(* Logix 5000 project; controller Seperator 1756-L85E rev 34.11; software revision 34.00; part 2 of 7 *)
(* tags used below, declared in another part *)
   Inp : BOOL;   // Alarm Condition Input 1=Alarm
   Cfg_Exists : BOOL;   // 1=Alarm configured to exist, 0=Does not exist, don't scan
   Cfg_ResetReqd : BOOL;   // 1=Latched Alarm, a Reset is required to clear this Alarm
   Cfg_AckReqd : BOOL;   // 1=Acknowledge required for this Alarm
   Cfg_AllowShelve : BOOL;   // 1=Allow Operator to Shelve this Alarm
   Cfg_AllowDisable : BOOL;   // 1=Allow Maintenance to Disable this Alarm
   Cfg_Severity : SINT;   // Alarm Severity: 1=Low, 2=Medium, 3=High, 4=Highest
   Cfg_AlmMinOnT : DINT;   // Minimum time Alm output stays on (sec)
   Cfg_MaxShelfT : INT;   // Auto unshelve after shelved this long (1..32767 minutes)
   PCfg_AllowExist : BOOL;   // 1=Alarm can be configured to exist, 0=other configs make alarm meaningless
   PCmd_Ack : BOOL;   // Program Command to Acknowledge alarm
   PCmd_Suppress : BOOL;   // Program Command to Suppress by Design (inhibits new alarm)
   PCmd_Unsuppress : BOOL;   // Program Command to Unsuppress (allows new alarm)
   PCmd_Unshelve : BOOL;   // Program Command to Unshelve (e.g., on shift change)
   OCmd_Ack : BOOL;   // Operator Command to Acknowledge alarm
   OCmd_Shelve : BOOL;   // Operator Command to Shelve Alarm (inhibits new alarm)
   OCmd_Unshelve : BOOL;   // Operator Command to Unshelve alarm (allows new alarm)
   Alm : ALIAS FOR Com_AE.0;   // Alarm output 1=In Alarm
   Ack : ALIAS FOR Com_AE.1;   // Alarm acknowledged status: 1=Ack rcvd
   Shelved : ALIAS FOR Com_AE.3;   // 1=Alarm has been Shelved by Operator (inhibits new alarm)
   Suppressed : ALIAS FOR Com_AE.6;   // 1=Alarm has been Suppressed by Program (inhibits new alarm)
   Disabled : ALIAS FOR Com_AE.9;   // 1=Alarm has been Disabled by Maintanance (inhibits new alarm)
   P_Alarm : BOOL;   // Unique Parameter Name for auto - discovery
   Wrk_Suppressed : BOOL;   // Internal Alarm Suppressed Status
   Com_AE : INT;   // Communication with HMI / Alarm/Event Server (see bit descriptions)
   Starting : SFC_STEP;
   Stopped : SFC_STEP;
   Stopping : SFC_STEP;
(* P_Alarm, continued *)

ROUTINE Prescan   (* ladder *)
// Clear "lurking" Commands
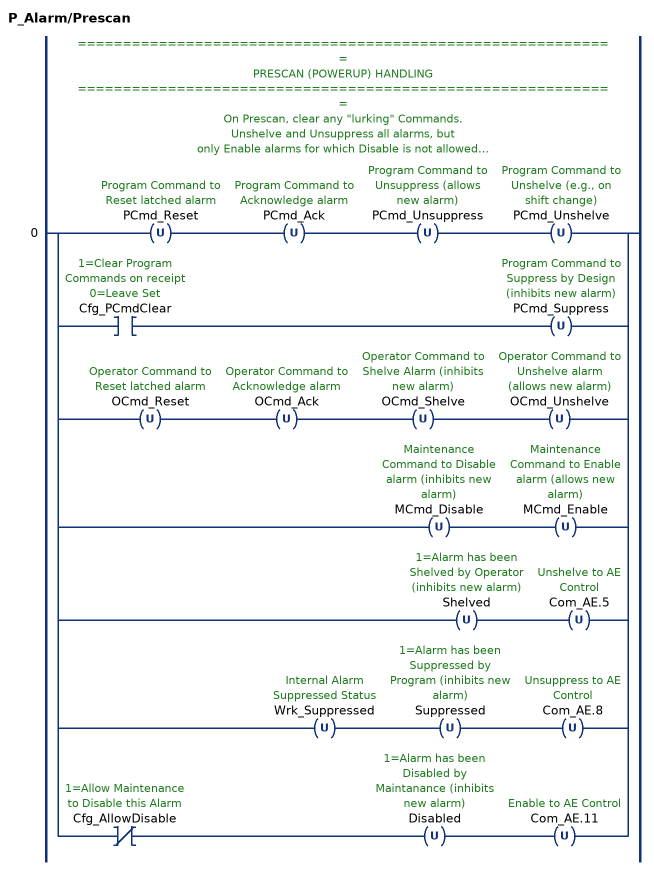
   // ============================================================
   // PRESCAN (POWERUP) HANDLING
   // ============================================================
   // On Prescan, clear any "lurking" Commands.
   // Unshelve and Unsuppress all alarms, but
   // only Enable alarms for which Disable is not allowed.
   // (Let Maintenance Disable persist through a power cycle...)
   // #####  V3.0-00  2013-06-30:  Added PCmd_Unshelve, AllowDisable, AllowShelve.  #####
   0: [OTU(PCmd_Reset) OTU(PCmd_Ack) OTU(PCmd_Unsuppress) OTU(PCmd_Unshelve) ,XIC(Cfg_PCmdClear) OTU(PCmd_Suppress) ,OTU(OCmd_Reset) OTU(OCmd_Ack) OTU(OCmd_Shelve) OTU(OCmd_Unshelve) ,OTU(MCmd_Disable) OTU(MCmd_Enable) ,OTU(Shelved) OTU(Com_AE.5) ,OTU(Wrk_Suppressed) OTU(Suppressed) OTU(Com_AE.8) ,XIO(Cfg_AllowDisable) OTU(Disabled) OTU(Com_AE.11) ];
END_ROUTINE
END_ADD_ON_INSTRUCTION

ADD_ON_INSTRUCTION P_Mode   (* revision 3.0 00 Release, vendor Rockwell Automation, ExecutePrescan, ExecuteEnableInFalse *)
// Mode
// Revision note:
// See Release Notes for Library version 3.0 for details on changes for this release. Containing objects MUST now expose OCmd_AcqLock and OCmd_Unlock. Made Operator Commands for going from Operator Locked to Program (unlocked) and Program (unlocked) to Operator Lock two-step processes.  Added Inf_Lib, Inf_Type.
// Help:
// Copyright © Rockwell Automation, Inc.  All Rights Reserved.
// This instruction provides selection of Mode (owner) for a Device level
// object  (from highest priority to lowest):
// *  No Mode (no owner, EnableIn is false)
// *  Hand (typically tracks hardwired control of device)
// *  Maint (Maintenance) (taken out of normal service for maintenance)
// *  Ovrd (Override) (typically used for process overrides)
// *  Prog  (Program) (automated control, and default if Cfg_ProgNorm = 1)
// *  Oper (Operator (manual control, and default if Cfg_ProgNorm = 0)
// (Program and Operator have the same priority.)
// The current mode is shown with Status bits and also as the primary
// Value for the instruction: an enumeration "Val" as follows:
//   0 = No Mode,
//   1 = Hand,
//   2 = Maintenance,
//   3 = Override,
//   4 = Program (Locked),
//   5 = Operator (Locked),
//   6 = Program (Unlocked, Oper default),
//   7 = Operator (Unlocked, Prog default),
//   8 = Program (Unlocked, = default),
//   9 = Operator (Unlocked, = default).
// When EnableIn is false, all ownership acquire/release and lock/unlock
// Commands are processed "behind the scenes", but the Mode is shown
// as "No Mode" (no owner).  When EnableIn becomes true, the Mode
// takes into account the Commands received -- in other words, the Mode
// becomes the one that would have been in effect had the EnableIn
// False / No Mode condition never occurred.
VAR_INPUT
   Inp_Hand : BOOL; {visible}   // 1=Acquire Hand (typ. hardwired local) Mode, 0=Release Hand Mode
   Inp_Ovrd : BOOL; {visible}   // 1=Acquire Override (higher priority program logic) Mode, 0=Release Override Mode
   Cfg_PCmdClear : BOOL := 1;   // 1=Clear Program Command on receipt; 0=Use Level-based (maintained) PCmds
   Cfg_OvrdOverLock : BOOL := 1;   // 1=Override supersedes Prog/Oper Lock, 0=don't override Lock
   Cfg_ProgDefault : BOOL;   // Default Mode: 1=Program Mode if no requests; 0=Operator Mode if no requests
   PCmd_Acq : BOOL;   // Program Command to Acquire Ownership (Oper to Prog)
   PCmd_Rel : BOOL;   // Program Command to Release Ownership (Prog to Oper)
   PCmd_Lock : BOOL;   // Program Command to Lock Mode in Prog
   PCmd_Unlock : BOOL;   // Program Command to Unlock Mode
   MCmd_Acq : BOOL;   // Maintenance Command to Acquire Ownership (Oper/Prog/Ovrd to Maint)
   MCmd_Rel : BOOL;   // Maintenance Command to Release Ownership (Maint to Oper/Prog/Ovrd)
   OCmd_AcqLock : BOOL;   // Operator Command to Acquire (Prog to Oper) / Lock Ownership
   OCmd_UnlockRel : BOOL;   // Operator Command to Unlock / Release (Oper to Prog) Ownership
END_VAR
VAR_OUTPUT
   Val : DINT; {access Read Only}   // Mode enum: 0=No, 1=H, 2=M, 3=!, 4=P Lock, 5=O Lock, 6=P (O Def), 7=O (P Def), 8=P (= Def), 9=O (= Def)
   Sts_Hand : BOOL; {access Read Only, visible}   // 1=Mode is Hand (supersedes Maint, Ovrd, Prog, Oper)
   Sts_Maint : BOOL; {access Read Only, visible}   // 1=Mode is Maintenance (supersedes Ovrd, Prog, Oper)
   Sts_Ovrd : BOOL; {access Read Only, visible}   // 1=Mode is Override (supersedes Prog, Oper)
   Sts_Prog : BOOL; {access Read Only, visible}   // 1=Mode is Program
   Sts_Oper : BOOL := 1; {access Read Only, visible}   // 1=Mode is Operator
   Sts_ProgOperLock : BOOL; {access Read Only, visible}   // 1=Program or Operator has requested Mode Lock
   Sts_ProgOperSel : BOOL; {access Read Only}   // Prog/Oper selection 1=Program, 0=Operator
   Sts_NoMode : BOOL; {access Read Only}   // 1=Mode is No Mode (no owner, disabled or not scanned)
   Rdy_MAcq : BOOL; {access Read Only}   // 1=Ready for MCmd_Acq, enable button
   Rdy_MRel : BOOL; {access Read Only}   // 1=Ready for MCmd_Rel, enable button
   Rdy_OAcq : BOOL; {access Read Only}   // 1=Ready for OCmd_AcqLock, enable Acquire (to Oper) button
   Rdy_OLock : BOOL; {access Read Only}   // 1=Ready for OCmd_AcqLock, enable Oper Lock button
   Rdy_OUnlock : BOOL; {access Read Only}   // 1=Ready for OCmd_UnlockRel, enable Oper Unlock button
   Rdy_ORel : BOOL; {access Read Only}   // 1=Ready for OCmd_UnlockRel, enable Release (to Prog) button
   P_Mode : BOOL;   // Unique Parameter Name for auto - discovery
END_VAR
VAR
   Wrk_Locked : BOOL; {access None}   // 1=Program/Operator Mode selection is Locked
   Wrk_Prog : BOOL; {access None}   // Internal Program (1) / Operator (0) Mode selection
   Wrk_Maint : BOOL; {access None}   // Internal Maintenance Mode
   Inf_Lib : STRING_12 := 'RA-BAS'; {access Read Only}   // Display Library for Faceplate call-up
   Inf_Type : STRING_16_UDT := 'P_Mode'; {access Read Only}   // Must contain AOI name, used for HMI and Information S/W
END_VAR

ROUTINE EnableInFalse   (* ladder *)
// Processes received Commands, but shows "NO mode" (no owner)
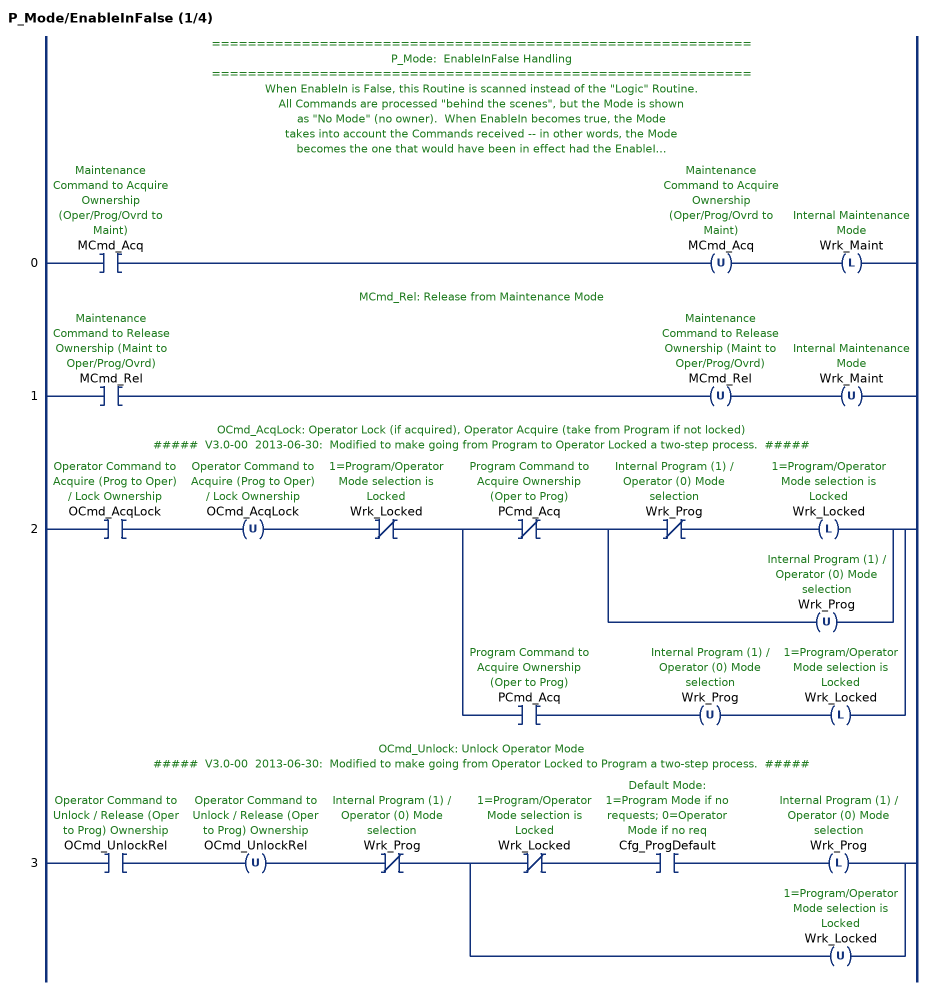
   // ============================================================
   // P_Mode:  EnableInFalse Handling
   // ============================================================
   // When EnableIn is False, this Routine is scanned instead of the "Logic" Routine.
   // All Commands are processed "behind the scenes", but the Mode is shown
   // as "No Mode" (no owner).  When EnableIn becomes true, the Mode
   // takes into account the Commands received -- in other words, the Mode
   // becomes the one that would have been in effect had the EnableIn
   // False / No Mode condition never occurred.
   // ============================================================
   // COMMAND HANDLING
   // ============================================================
   // NOTE:  These rungs MUST be in the order given to meet the following
   // multiple-actions-at-the-same-time scenarios:
   // * Maintenance Release beats Maintenance Acquire
   // * Program Release beats Program Acquire
   // * Program Unlock beats Program Lock
   // * Operator Unlock beats Operator Acquire and Lock (results in Oper Unlocked)
   // * Operator Acquire/Lock must come after Program Unlock
   // * Program Acquire must come after Operator Unlock
   // ============================================================
   // MCmd_Acq: Acquire for Maintenance Mode
   0: XIC(MCmd_Acq)OTU(MCmd_Acq)OTL(Wrk_Maint);
   // MCmd_Rel: Release from Maintenance Mode
   1: XIC(MCmd_Rel)OTU(MCmd_Rel)OTU(Wrk_Maint);
   // OCmd_AcqLock: Operator Lock (if acquired), Operator Acquire (take from Program if not locked)
   // #####  V3.0-00  2013-06-30:  Modified to make going from Program to Operator Locked a two-step process.  #####
   2: XIC(OCmd_AcqLock)OTU(OCmd_AcqLock)XIO(Wrk_Locked)[XIO(PCmd_Acq) [XIO(Wrk_Prog) OTL(Wrk_Locked) ,OTU(Wrk_Prog) ] ,XIC(PCmd_Acq) OTU(Wrk_Prog) OTL(Wrk_Locked) ];
   // OCmd_Unlock: Unlock Operator Mode
   // #####  V3.0-00  2013-06-30:  Modified to make going from Operator Locked to Program a two-step process.  #####
   3: XIC(OCmd_UnlockRel)OTU(OCmd_UnlockRel)XIO(Wrk_Prog)[XIO(Wrk_Locked) XIC(Cfg_ProgDefault) OTL(Wrk_Prog) ,OTU(Wrk_Locked) ];
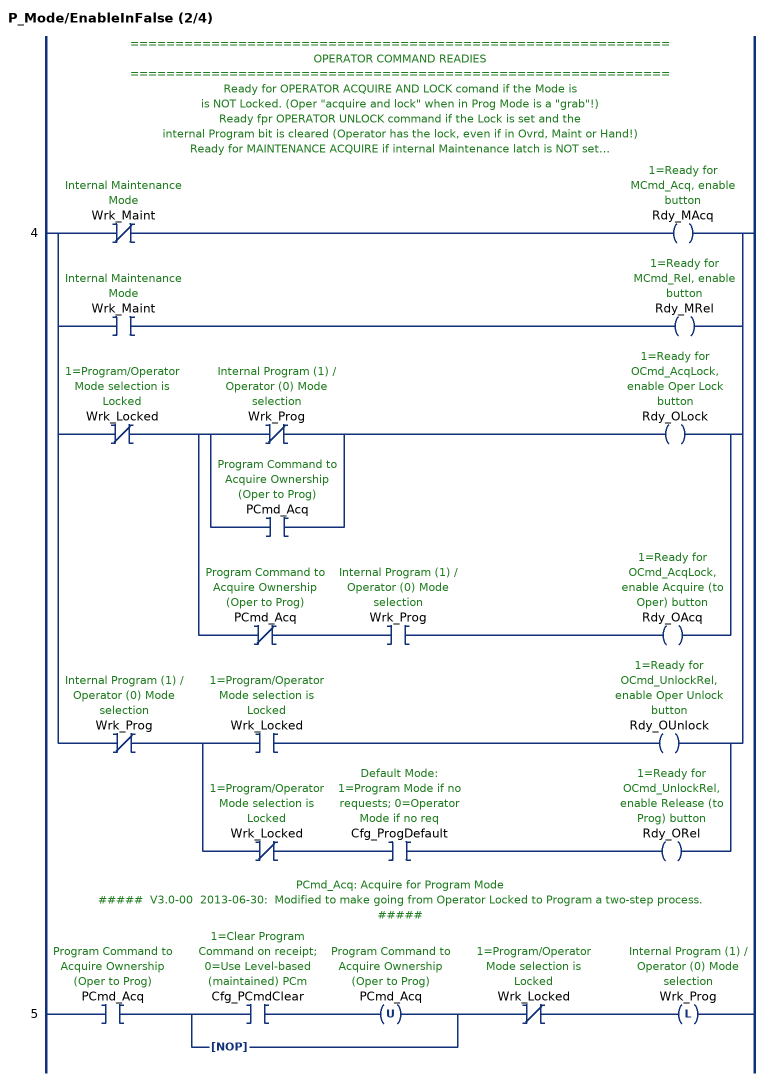
   // ============================================================
   // OPERATOR COMMAND READIES
   // ============================================================
   // Ready for OPERATOR ACQUIRE AND LOCK comand if the Mode is
   //  is NOT Locked. (Oper "acquire and lock" when in Prog Mode is a "grab"!)
   // Ready fpr OPERATOR UNLOCK command if the Lock is set and the
   // internal Program bit is cleared (Operator has the lock, even if in Ovrd, Maint or Hand!)
   // Ready for MAINTENANCE ACQUIRE if internal Maintenance latch is NOT set.
   // Ready for MAINTENANCE RELEASE if internal Maintenance latch IS set.
   // #####  V3.0-00  2013-06-30:  Modified Rdy_Unlock for two-step Operator Locked to Program process.  #####
   4: [XIO(Wrk_Maint) OTE(Rdy_MAcq) ,XIC(Wrk_Maint) OTE(Rdy_MRel) ,XIO(Wrk_Locked) [[XIO(Wrk_Prog) ,XIC(PCmd_Acq) ] OTE(Rdy_OLock) ,XIO(PCmd_Acq) XIC(Wrk_Prog) OTE(Rdy_OAcq) ] ,XIO(Wrk_Prog) [XIC(Wrk_Locked) OTE(Rdy_OUnlock) ,XIO(Wrk_Locked) XIC(Cfg_ProgDefault) OTE(Rdy_ORel) ] ];
   // PCmd_Acq: Acquire for Program Mode
   // #####  V3.0-00  2013-06-30:  Modified to make going from Operator Locked to Program a two-step process.  #####
   5: XIC(PCmd_Acq)[XIC(Cfg_PCmdClear) OTU(PCmd_Acq) ,NOP() ]XIO(Wrk_Locked)OTL(Wrk_Prog);
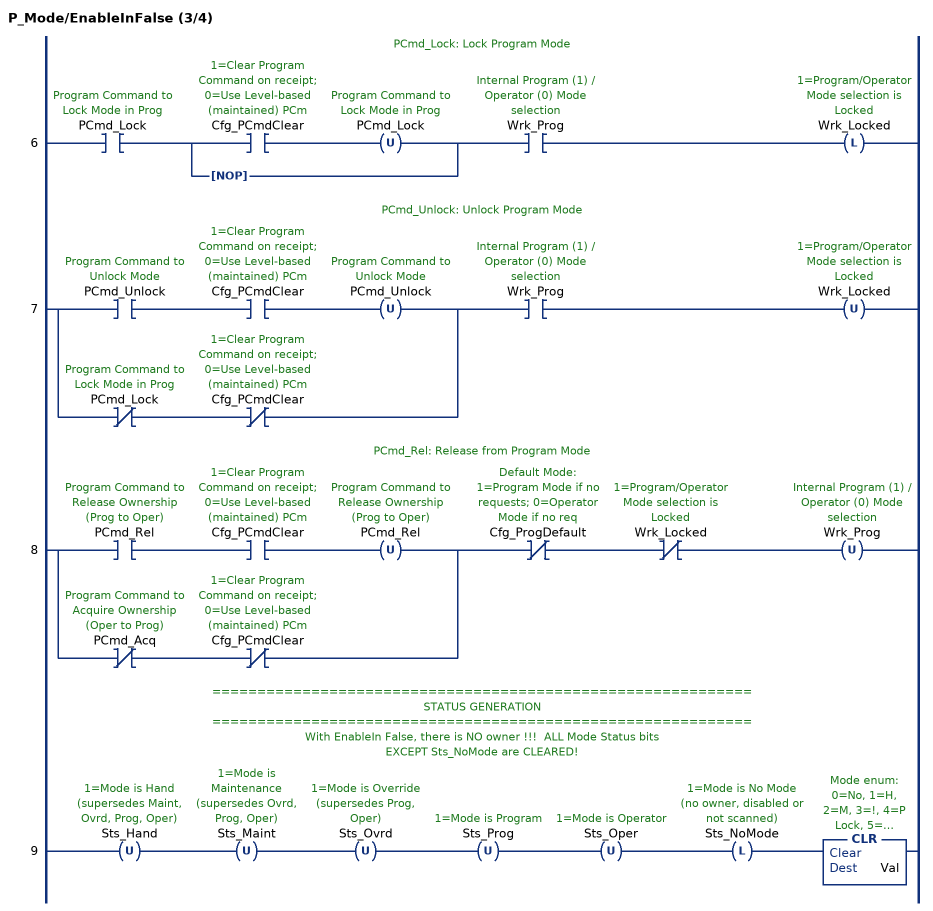
   // PCmd_Lock: Lock Program Mode
   6: XIC(PCmd_Lock)[XIC(Cfg_PCmdClear) OTU(PCmd_Lock) ,NOP() ]XIC(Wrk_Prog)OTL(Wrk_Locked);
   // PCmd_Unlock: Unlock Program Mode
   7: [XIC(PCmd_Unlock) XIC(Cfg_PCmdClear) OTU(PCmd_Unlock) ,XIO(PCmd_Lock) XIO(Cfg_PCmdClear) ]XIC(Wrk_Prog)OTU(Wrk_Locked);
   // PCmd_Rel: Release from Program Mode
   8: [XIC(PCmd_Rel) XIC(Cfg_PCmdClear) OTU(PCmd_Rel) ,XIO(PCmd_Acq) XIO(Cfg_PCmdClear) ]XIO(Cfg_ProgDefault)XIO(Wrk_Locked)OTU(Wrk_Prog);
   // ============================================================
   // STATUS GENERATION
   // ============================================================
   // With EnableIn False, there is NO owner !!!  ALL Mode Status bits
   // EXCEPT Sts_NoMode are CLEARED!
   9: OTU(Sts_Hand)OTU(Sts_Maint)OTU(Sts_Ovrd)OTU(Sts_Prog)OTU(Sts_Oper)OTL(Sts_NoMode)CLR(Val);
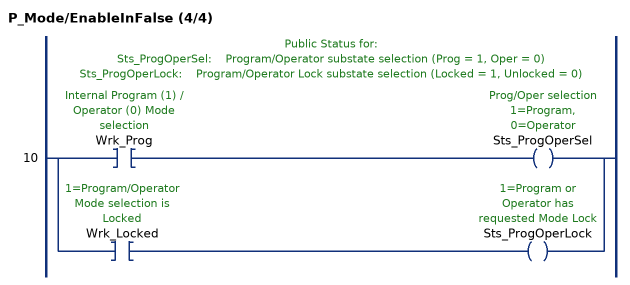
   // Public Status for:
   // Sts_ProgOperSel:    Program/Operator substate selection (Prog = 1, Oper = 0)
   // Sts_ProgOperLock:    Program/Operator Lock substate selection (Locked = 1, Unlocked = 0)
   10: [XIC(Wrk_Prog) OTE(Sts_ProgOperSel) ,XIC(Wrk_Locked) OTE(Sts_ProgOperLock) ];
END_ROUTINE

ROUTINE Logic   (* ladder *)
// Selects Modes (Hand, Maint, Ovrd, Oper, Prog) based on Inputs and Commands
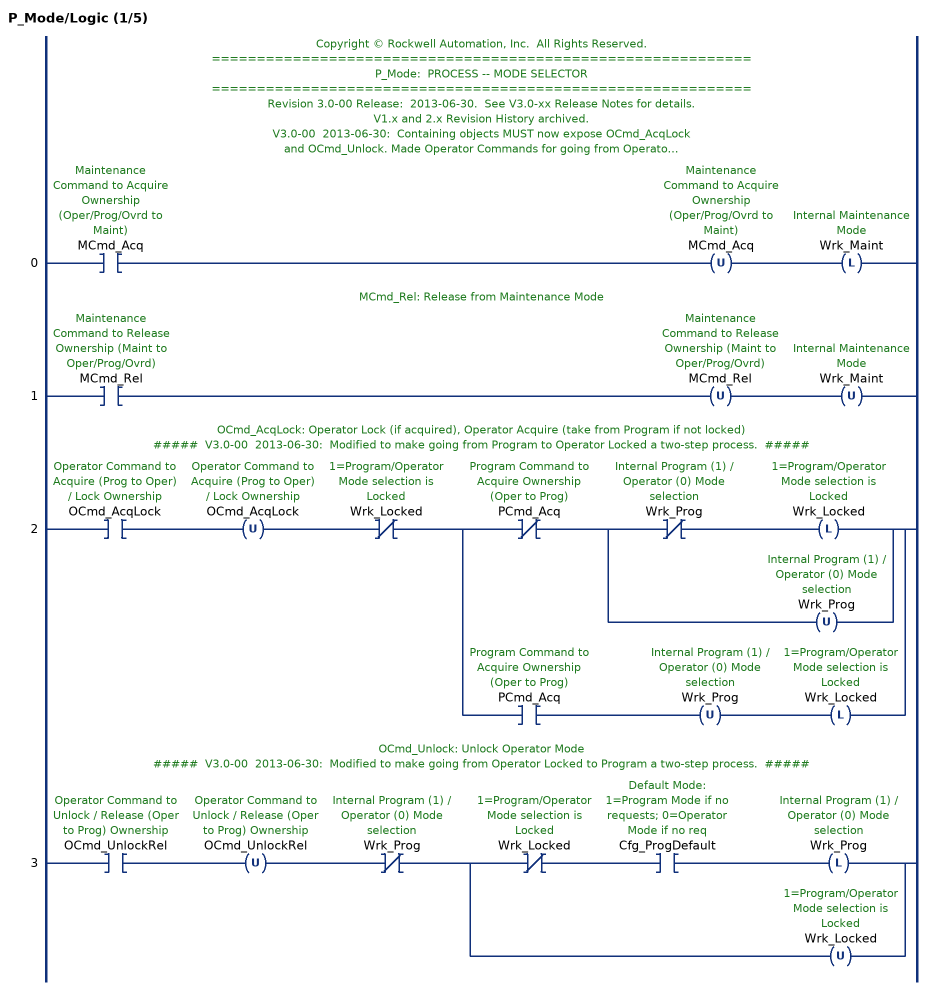
   // Copyright © Rockwell Automation, Inc.  All Rights Reserved.
   // ============================================================
   // P_Mode:  PROCESS -- MODE SELECTOR
   // ============================================================
   // Revision 3.0-00 Release:  2013-06-30.  See V3.0-xx Release Notes for details.
   // V1.x and 2.x Revision History archived.
   // V3.0-00  2013-06-30:  Containing objects MUST now expose OCmd_AcqLock
   // and OCmd_Unlock. Made Operator Commands for going from Operator
   // Locked to Program (unlocked) and Program (unlocked) to Operator
   // Lock two-step processes.  Added Inf_Lib, Inf_Type.
   // ============================================================
   // This instruction provides selection of Mode (owner) for a Device level
   // object  (from highest priority to lowest):
   // * NO Mode (EnableIn is false)
   // *  Hand (typically tracks hardwired control of device)
   // *  Maint (Maintenance) (taken out of normal service for maintenance)
   // *  Ovrd (Override) (typically used for process overrides)
   // *  Prog  (Program) (automated control, and default if Cfg_ProgNorm = 1)
   // *  Oper (Operator (manual control, and default if Cfg_ProgNorm = 0)
   // The current mode is shown with Status bits and also as the
   // primary Value for the instruction: an enumeration as follows:
   // 0 = No Mode, 1 = Hand, 2 = Maintenance, 3 = Override,
   // 4 = Program (Locked), 5 = Operator (Locked),
   // 6 = Program (Unlocked, Oper default), 7 = Operator (Unlocked, Prog default),
   // 8 = Program (Unlocked, Prog default), 9 = Operator (Unlocked, Oper default).
   // ============================================================
   // COMMAND HANDLING
   // ============================================================
   // NOTE:  These rungs MUST be in the order given to meet the following
   // multiple-actions-at-the-same-time scenarios:
   // * Maintenance Release beats Maintenance Acquire
   // * Program Release beats Program Acquire
   // * Program Unlock beats Program Lock
   // * Operator Unlock beats Operator Acquire / Lock (results in Oper Unlocked)
   // * Program Acquire must come after Operator Unlock
   // If Cfg_ProgDefault = 1, the Mode defaults to Program
   // (instead of Operator) if all other Modes release their requests.
   // ============================================================
   // MCmd_Acq: Acquire for Maintenance Mode
   0: XIC(MCmd_Acq)OTU(MCmd_Acq)OTL(Wrk_Maint);
   // MCmd_Rel: Release from Maintenance Mode
   1: XIC(MCmd_Rel)OTU(MCmd_Rel)OTU(Wrk_Maint);
   // OCmd_AcqLock: Operator Lock (if acquired), Operator Acquire (take from Program if not locked)
   // #####  V3.0-00  2013-06-30:  Modified to make going from Program to Operator Locked a two-step process.  #####
   2: XIC(OCmd_AcqLock)OTU(OCmd_AcqLock)XIO(Wrk_Locked)[XIO(PCmd_Acq) [XIO(Wrk_Prog) OTL(Wrk_Locked) ,OTU(Wrk_Prog) ] ,XIC(PCmd_Acq) OTU(Wrk_Prog) OTL(Wrk_Locked) ];
   // OCmd_Unlock: Unlock Operator Mode
   // #####  V3.0-00  2013-06-30:  Modified to make going from Operator Locked to Program a two-step process.  #####
   3: XIC(OCmd_UnlockRel)OTU(OCmd_UnlockRel)XIO(Wrk_Prog)[XIO(Wrk_Locked) XIC(Cfg_ProgDefault) OTL(Wrk_Prog) ,OTU(Wrk_Locked) ];
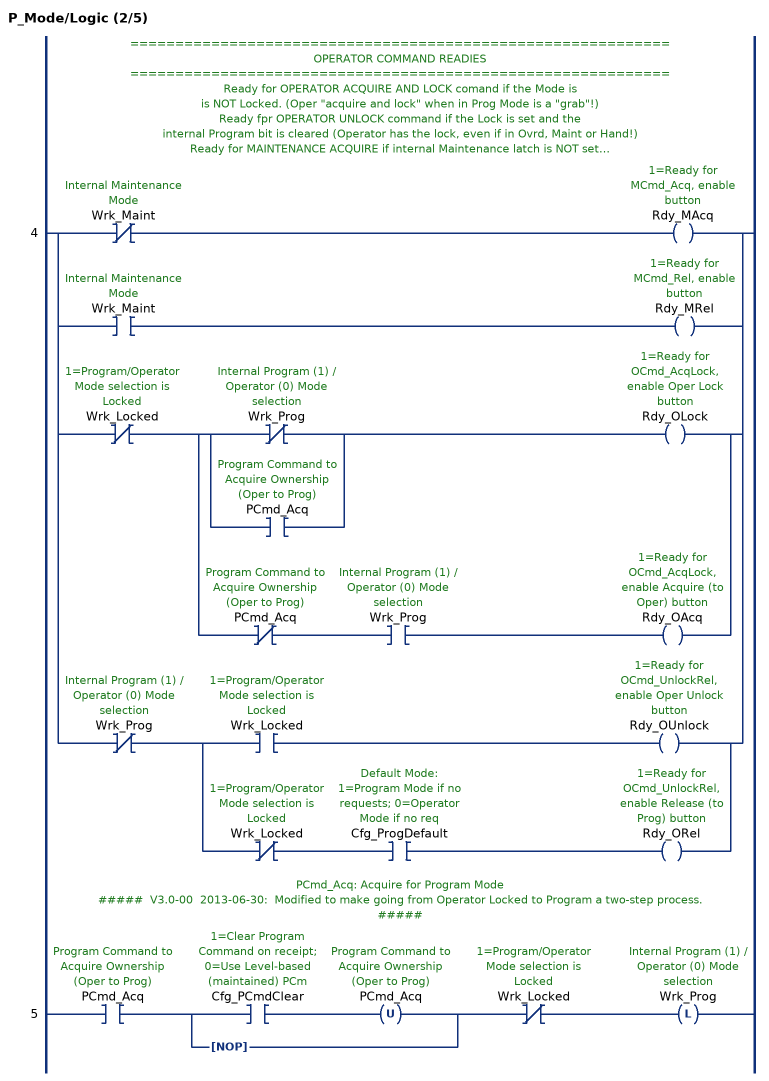
   // ============================================================
   // OPERATOR COMMAND READIES
   // ============================================================
   // Ready for OPERATOR ACQUIRE AND LOCK comand if the Mode is
   //  is NOT Locked. (Oper "acquire and lock" when in Prog Mode is a "grab"!)
   // Ready fpr OPERATOR UNLOCK command if the Lock is set and the
   // internal Program bit is cleared (Operator has the lock, even if in Ovrd, Maint or Hand!)
   // Ready for MAINTENANCE ACQUIRE if internal Maintenance latch is NOT set.
   // Ready for MAINTENANCE RELEASE if internal Maintenance latch IS set.
   // #####  V3.0-00  2013-06-30:  Modified Rdy_Unlock for two-step Operator Locked to Program process.  #####
   4: [XIO(Wrk_Maint) OTE(Rdy_MAcq) ,XIC(Wrk_Maint) OTE(Rdy_MRel) ,XIO(Wrk_Locked) [[XIO(Wrk_Prog) ,XIC(PCmd_Acq) ] OTE(Rdy_OLock) ,XIO(PCmd_Acq) XIC(Wrk_Prog) OTE(Rdy_OAcq) ] ,XIO(Wrk_Prog) [XIC(Wrk_Locked) OTE(Rdy_OUnlock) ,XIO(Wrk_Locked) XIC(Cfg_ProgDefault) OTE(Rdy_ORel) ] ];
   // PCmd_Acq: Acquire for Program Mode
   // #####  V3.0-00  2013-06-30:  Modified to make going from Operator Locked to Program a two-step process.  #####
   5: XIC(PCmd_Acq)[XIC(Cfg_PCmdClear) OTU(PCmd_Acq) ,NOP() ]XIO(Wrk_Locked)OTL(Wrk_Prog);
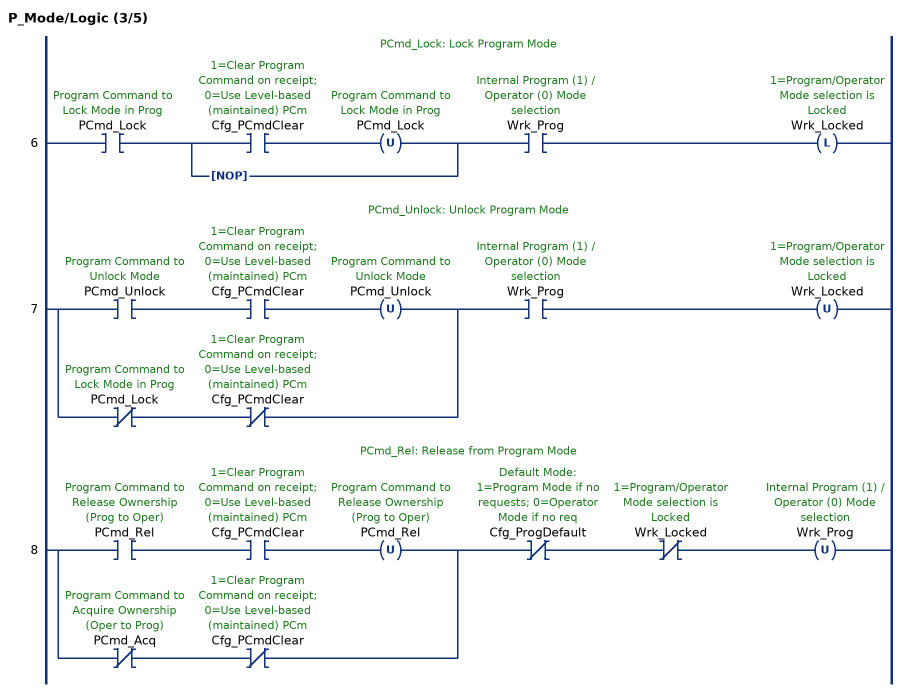
   // PCmd_Lock: Lock Program Mode
   6: XIC(PCmd_Lock)[XIC(Cfg_PCmdClear) OTU(PCmd_Lock) ,NOP() ]XIC(Wrk_Prog)OTL(Wrk_Locked);
   // PCmd_Unlock: Unlock Program Mode
   7: [XIC(PCmd_Unlock) XIC(Cfg_PCmdClear) OTU(PCmd_Unlock) ,XIO(PCmd_Lock) XIO(Cfg_PCmdClear) ]XIC(Wrk_Prog)OTU(Wrk_Locked);
   // PCmd_Rel: Release from Program Mode
   8: [XIC(PCmd_Rel) XIC(Cfg_PCmdClear) OTU(PCmd_Rel) ,XIO(PCmd_Acq) XIO(Cfg_PCmdClear) ]XIO(Cfg_ProgDefault)XIO(Wrk_Locked)OTU(Wrk_Prog);
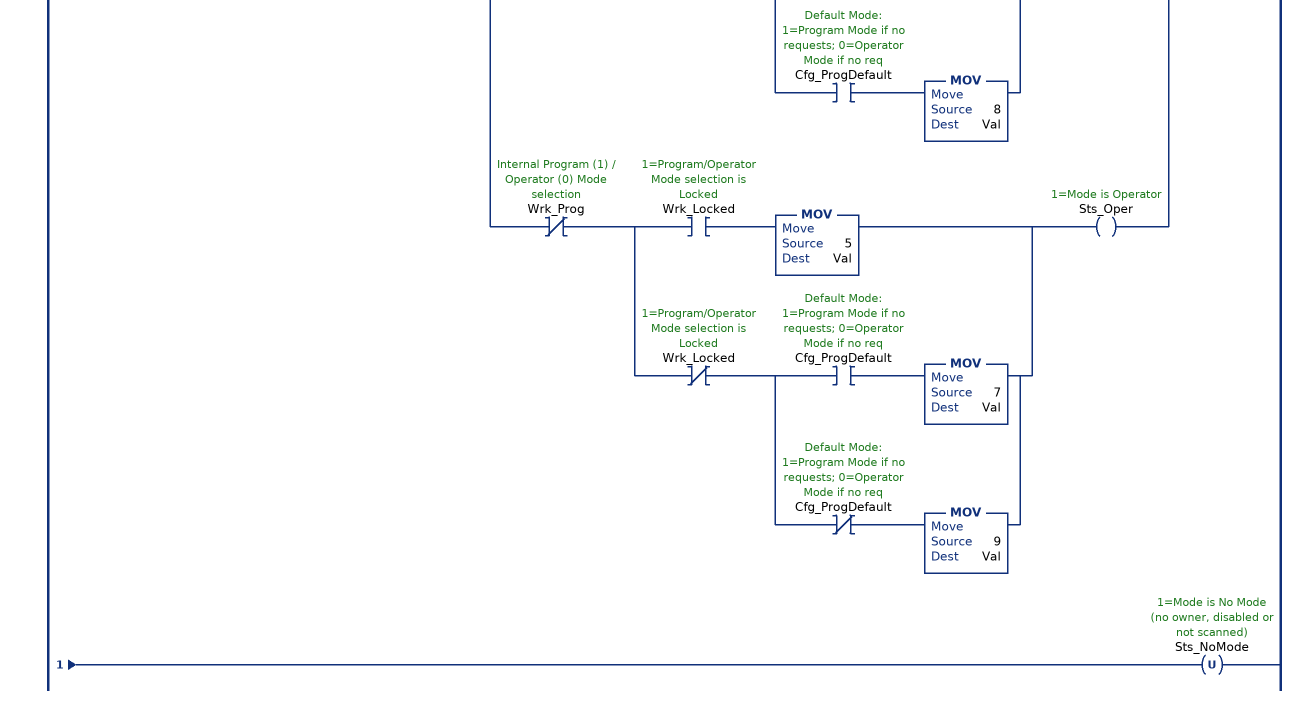
   // ============================================================
   // STATUS GENERATION
   // ============================================================
   // This rung determines the Mode based on the states of the inputs and internal working bits.
   // The logic here does the vast mahority of the implementation of the Mode selection rules.
   // Between the internal working bits used above and the rules implemented here,
   // outside objects cannot manipulate the state of this object by setting/clearing its Status bits.
   // Public Status is generated for:
   // *  Hand Mode
   // *  Maintenance Mode
   // *  Override Mode
   // *  Program Mode
   // *  Operator Mode
   // *  No Mode (none of the above)
   9: [XIC(Inp_Hand) OTE(Sts_Hand) MOV(1,Val) ,XIO(Inp_Hand) [XIC(Wrk_Maint) OTE(Sts_Maint) MOV(2,Val) ,XIO(Wrk_Maint) [XIC(Inp_Ovrd) [XIO(Wrk_Locked) ,XIC(Cfg_OvrdOverLock) ,XIC(Sts_Ovrd) ] OTE(Sts_Ovrd) MOV(3,Val) ,XIO(Sts_Ovrd) [XIC(Wrk_Prog) [XIC(Wrk_Locked) MOV(4,Val) ,XIO(Wrk_Locked) [XIO(Cfg_ProgDefault) MOV(6,Val) ,XIC(Cfg_ProgDefault) MOV(8,Val) ] ] OTE(Sts_Prog) ,XIO(Wrk_Prog) [XIC(Wrk_Locked) MOV(5,Val) ,XIO(Wrk_Locked) [XIC(Cfg_ProgDefault) MOV(7,Val) ,XIO(Cfg_ProgDefault) MOV(9,Val) ] ] OTE(Sts_Oper) ] ] ] ]OTU(Sts_NoMode);
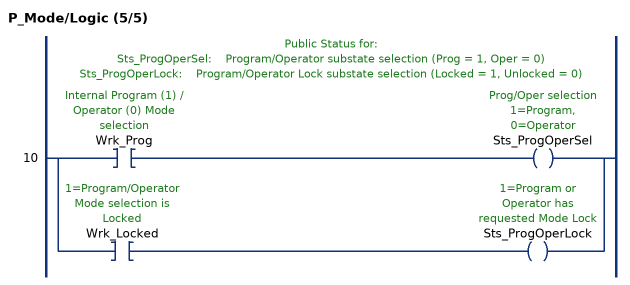
   // Public Status for:
   // Sts_ProgOperSel:    Program/Operator substate selection (Prog = 1, Oper = 0)
   // Sts_ProgOperLock:    Program/Operator Lock substate selection (Locked = 1, Unlocked = 0)
   10: [XIC(Wrk_Prog) OTE(Sts_ProgOperSel) ,XIC(Wrk_Locked) OTE(Sts_ProgOperLock) ];
END_ROUTINE

ROUTINE Prescan   (* ladder *)
// Clear "lurking" Commands
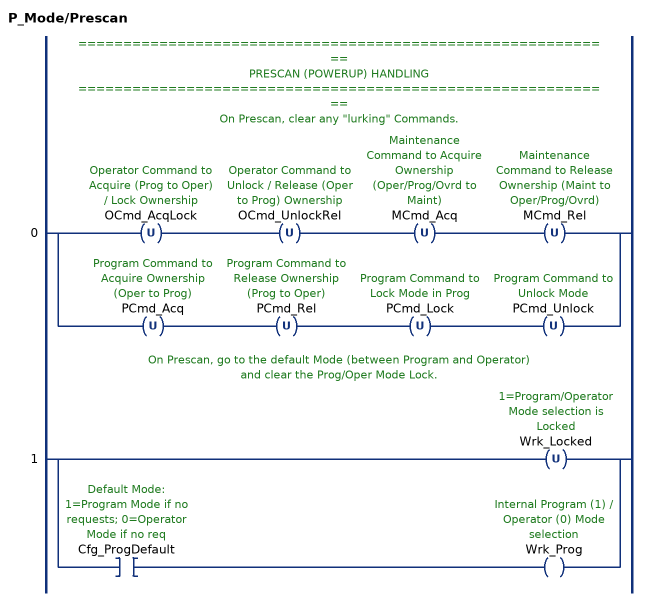
   // ============================================================
   // PRESCAN (POWERUP) HANDLING
   // ============================================================
   // On Prescan, clear any "lurking" Commands.
   0: [OTU(OCmd_AcqLock) OTU(OCmd_UnlockRel) OTU(MCmd_Acq) OTU(MCmd_Rel) ,OTU(PCmd_Acq) OTU(PCmd_Rel) OTU(PCmd_Lock) OTU(PCmd_Unlock) ];
   // On Prescan, go to the default Mode (between Program and Operator)
   // and clear the Prog/Oper Mode Lock.
   1: [OTU(Wrk_Locked) ,XIC(Cfg_ProgDefault) OTE(Wrk_Prog) ];
END_ROUTINE
END_ADD_ON_INSTRUCTION

ADD_ON_INSTRUCTION P_Motor   (* revision 3.0 04 Release, vendor Rockwell Automation, ExecutePrescan, ExecuteEnableInFalse *)
// Single Speed Motor
// Revision note:
// See Release Notes for Library version 3.0 for details on changes for this release. Corrected Parameter descriptions and default configuration values for alarms only.
// Help:
// Copyright © Rockwell Automation, Inc.  All Rights Reserved.
// This Instruction controls and monitors a single-speed motor
// (FVNR, soft-start, etc.) and provides:
// *  Monitoring of run feedback, display of actual motor status
// *  Detection of Failure to Start, Failure to Stop
// *  Monitoring of a Permissive condition to allow starting
// *  Monitoring of an Interlock condition to stop / prevent starting
// *  Simulation, providing feedback of a working motor while disabling outputs
// *  Monitoring of I/O communication faults
// *  Alarms for Fail to Start, Fail to Stop, Interlock Trip, I/O Fault
// *  Options to shed (stop motor) on Fail to Start or I/O Fault
// *  Operation in Hand, Maintenance, Override, Program and Operator Modes
// *  Option to automatically reset faults and alarms when operator commands
//      motor to start or stop
// *  Supports HMI "breadcrumbs" for Alarm Inhibited, Bad Configuration,
//      Not Ready, Maintenance Bypass Active
// *  "Available" status for use by automation logic to know whether motor
//      can be controlled by other objects.
// Modes are provided by a P_Mode AOI instance.
// Alarms are provided by P_Alarm AOI instances.
// Modes of operation: Operator, Program, Override, Maintenance, Hand
VAR_INPUT
   Inp_RunFdbk : BOOL; {visible}   // Input Signal: RUN feedback from motor
   Inp_PermOK : BOOL := 1; {visible}   // 1=Permissives OK, motor can start
   Inp_NBPermOK : BOOL := 1; {visible}   // 1=Non-Bypassable Permissives OK, motor can start
   Inp_IntlkOK : BOOL := 1; {visible}   // 1=Interlocks OK, motor can start/run
   Inp_NBIntlkOK : BOOL := 1; {visible}   // 1=Non-Bypassable Interlocks OK, motor can start/run
   Inp_IOFault : BOOL;   // Input Communication Status 0=OK, 1=fail
   Inp_Sim : BOOL;   // 1=Simulate working motor; 0=Start/Stop/ Monitor actual motor
   Inp_Hand : ALIAS FOR Mode.Inp_Hand;
   Inp_Ovrd : ALIAS FOR Mode.Inp_Ovrd;
   Inp_OvrdCmd : DINT;   // Override Mode Command: 0=None, 1=Stop, 2=Start
   Inp_Reset : BOOL;   // 1=Reset all fault conditions and latched Alarms
   Cfg_HasRunFdbk : BOOL;   // 1=Motor provides run feedback
   Cfg_UseRunFdbk : BOOL;   // 1=Motor run feedback should be used for failure checking
   Cfg_AllowLocal : BOOL;   // 1=Allow Local Start/Stop without alarm, 0=Start/Stop from HMI/prog only
   Cfg_HasPermObj : BOOL;   // 1=Enable navigation to permissive object
   Cfg_HasIntlkObj : BOOL;   // 1=Enable navigation to interlock object
   Cfg_HasResInhObj : BOOL;   // 1=Enable navigation to restart inhibit object
   Cfg_HasRunTimeObj : BOOL;   // 1=Enable navigation to run time object
   Cfg_HasOvldObj : BOOL;   // 1=Enable navigation to overload object
   Cfg_PCmdClear : ALIAS FOR Mode.Cfg_PCmdClear;
   Cfg_ProgDefault : ALIAS FOR Mode.Cfg_ProgDefault;
   Cfg_OperStopPrio : BOOL;   // 1=OCmd_Stop available in any mode, 0=OCmd_Stop only in Oper, Maint modes.
   Cfg_OCmdResets : BOOL;   // 1=New Oper motor cmd. resets fault, 0=reset req'd to clear fault
   Cfg_OvrdPermIntlk : BOOL;   // 1=Override ignores Bypassable Perm/ Intlk; 0=always use Perm/Intlk
   Cfg_ShedOnFailToStart : BOOL := 1;   // 1=Stop Motor and Alarm on Fail to Start; 0=Alarm only on Fail to Start
   Cfg_ShedOnIOFault : BOOL := 1;   // 1=Stop Motor and Alarm on I/O Fault; 0=Alarm only on I/O Fault
   Cfg_HasFailToStartAlm : ALIAS FOR FailToStart.Cfg_Exists;   // 1=Fail to Start Alarm exists and will be checked
   Cfg_HasFailToStopAlm : ALIAS FOR FailToStop.Cfg_Exists;   // 1=Fail to Stop Alarm exists and will be checked
   Cfg_HasIntlkTripAlm : ALIAS FOR IntlkTrip.Cfg_Exists;   // 1=Interlock Trip Alarm exists and will be checked
   Cfg_HasIOFaultAlm : ALIAS FOR IOFault.Cfg_Exists;   // 1=I/O Fault Alarm exists and will be checked
   Cfg_FailToStartResetReqd : ALIAS FOR FailToStart.Cfg_ResetReqd;   // 1=Reset required to clear Fail to Start Alarm
   Cfg_FailToStopResetReqd : ALIAS FOR FailToStop.Cfg_ResetReqd;   // 1=Reset required to clear Fail to Stop Alarm
   Cfg_IntlkTripResetReqd : ALIAS FOR IntlkTrip.Cfg_ResetReqd;   // 1=Reset required to clear Interlock Trip Alarm
   Cfg_IOFaultResetReqd : ALIAS FOR IOFault.Cfg_ResetReqd;   // 1=Reset required to clear I/O Fault Alarm
   Cfg_FailToStartAckReqd : ALIAS FOR FailToStart.Cfg_AckReqd;   // 1=Acknowledge required for Fail to Start Alarm
   Cfg_FailToStopAckReqd : ALIAS FOR FailToStop.Cfg_AckReqd;   // 1=Acknowledge required for Fail to Stop Alarm
   Cfg_IntlkTripAckReqd : ALIAS FOR IntlkTrip.Cfg_AckReqd;   // 1=Acknowledge required for Interlock Trip Alarm
   Cfg_IOFaultAckReqd : ALIAS FOR IOFault.Cfg_AckReqd;   // 1=Acknowledge required for I/O Fault Alarm
   Cfg_FailToStartSeverity : ALIAS FOR FailToStart.Cfg_Severity;   // Fail To Start Alarm Severity: 1=low, 2=medium, 3=high, 4=highest
   Cfg_FailToStopSeverity : ALIAS FOR FailToStop.Cfg_Severity;   // Fail To Stop Alarm Severity: 1=low, 2=medium, 3=high, 4=highest
   Cfg_IntlkTripSeverity : ALIAS FOR IntlkTrip.Cfg_Severity;   // Interlock Trip Alarm Severity: 1=low, 2=medium, 3=high, 4=highest
   Cfg_IOFaultSeverity : ALIAS FOR IOFault.Cfg_Severity;   // I/O Fault Alarm Severity: 1=low, 2=medium, 3=high, 4=highest
   Cfg_SimFdbkT : DINT := 2;   // Feedback delay in Simulation (sec)
   Cfg_FailToStartT : DINT := 10;   // Time after Start for running feedback before Fault (sec)
   Cfg_FailToStopT : DINT := 10;   // Time after Stop for stopped feedback (=0) before Fault (sec)
   PSet_Owner : DINT;   // Program Owner Request ID (non-zero) or Release (zero)
   PCmd_Start : BOOL;   // Program Command to Start Motor
   PCmd_Stop : BOOL;   // Program Command to Stop Motor
   PCmd_Acq : ALIAS FOR Mode.PCmd_Acq;
   PCmd_Rel : ALIAS FOR Mode.PCmd_Rel;
   PCmd_Lock : ALIAS FOR Mode.PCmd_Lock;
   PCmd_Unlock : ALIAS FOR Mode.PCmd_Unlock;
   PCmd_Reset : BOOL;   // Program Command to Reset all Alarms requiring Reset
   PCmd_FailToStartAck : ALIAS FOR FailToStart.PCmd_Ack;   // Program Command to Acknowledge Fail to Start Alarm
   PCmd_FailToStartSuppress : ALIAS FOR FailToStart.PCmd_Suppress;   // Program Command to Suppress Fail to Start Alarm
   PCmd_FailToStartUnsuppress : ALIAS FOR FailToStart.PCmd_Unsuppress;   // Program Command to Unsuppress Fail to Start Alarm
   PCmd_FailToStartUnshelve : ALIAS FOR FailToStart.PCmd_Unshelve;   // Program Command to Unshelve Fail to Start Alarm
   PCmd_FailToStopAck : ALIAS FOR FailToStop.PCmd_Ack;   // Program Command to Acknowledge Fail to Stop Alarm
   PCmd_FailToStopSuppress : ALIAS FOR FailToStop.PCmd_Suppress;   // Program Command to Suppress Fail to Stop Alarm
   PCmd_FailToStopUnsuppress : ALIAS FOR FailToStop.PCmd_Unsuppress;   // Program Command to Unsuppress Fail to Stop Alarm
   PCmd_FailToStopUnshelve : ALIAS FOR FailToStop.PCmd_Unshelve;   // Program Comnmand to Unshelve Fail to Stop Alarm
   PCmd_IntlkTripAck : ALIAS FOR IntlkTrip.PCmd_Ack;   // Program Command to Acknowledge Interlock Trip Alarm